(* CODESYS project codesys_webvisu_opcua.project

Project tree, tasks and I/O mapping:
  Device : CODESYS Control for Raspberry Pi SL, CODESYS GmbH, order no. 2302000009, version 4.8.0.0
    application app
      libraries: Standard, 3.5.18.0 (System); Memory, * (3S - Smart Software Solutions GmbH); Util, 3.5.19.0 (System); CmpSysEthernet, 3.4.3.0 (3S - Smart Software Solutions GmbH); VisuDialogs, * (System); CAA Callback Extern, 3.5.17.0 (CAA Technical Workgroup); SysTypes Interfaces, 3.5.2.0 (System); SysMem, 3.5.17.0 (System); CmpErrors Interfaces, * (System); CAA SerialCom, 3.5.17.0 (CAA Technical Workgroup); SysSocket, 3.5.19.0 (System)
      task MainTask (cyclic, interval 4 ms, priority 0) calls MAIN
      task VISU_TASK (cyclic, interval 100 ms, priority 31) calls VisuElems.Visu_Prg
      program MAIN [ST]
      Symbols
      visualisation VISU
      Kommunikationsverwalter
        OPC_UA_Symbols
          Informationsmodell
      function block FB_DEMO [ST]: add2
    SoftMotion General Axis Pool
      x_axis : SM_Drive_Virtual, 3S - Smart Software Solutions GmbH, order no. 1805, version 4.0.0.0
          settings: wDriveID = 0; fSWMaxVelocity = 100000; fSWMaxAcceleration = 100000; fSWMaxDeceleration = 100000; fRampJerk = 1e7; fSWLimitPositive = 3000; fSWLimitNegative = -500; fSWLimitDeceleration = 0.0; fSWErrorMaxDistance = 0.0
      y_axis : SM_Drive_Virtual, 3S - Smart Software Solutions GmbH, order no. 1805, version 4.0.0.0
          settings: fSWMaxVelocity = 100000; fSWMaxAcceleration = 100000; fSWMaxDeceleration = 100000; fRampJerk = 1e7; fSWLimitPositive = 3000; fSWLimitNegative = -3000; fSWLimitDeceleration = 0.0; fSWErrorMaxDistance = 0.0
      z_axis : SM_Drive_Virtual, 3S - Smart Software Solutions GmbH, order no. 1805, version 4.0.0.0
          settings: wDriveID = 2; fSWMaxVelocity = 100000; fSWMaxAcceleration = 100000; fSWMaxDeceleration = 100000; fRampJerk = 1e7; fSWLimitPositive = 100; fSWLimitNegative = -1000; fSWLimitDeceleration = 0.0; fSWErrorMaxDistance = 0.0
      a_axis : SM_Drive_Virtual, 3S - Smart Software Solutions GmbH, order no. 1805, version 4.0.0.0
          settings: wDriveID = 3; fSWMaxVelocity = 100000; fSWMaxAcceleration = 100000; fSWMaxDeceleration = 100000; fRampJerk = 1e7; fSWLimitPositive = 360; fSWLimitNegative = -360; fSWLimitDeceleration = 0.0; fSWErrorMaxDistance = 0.0
      r_axis : SM_Drive_Virtual, 3S - Smart Software Solutions GmbH, order no. 1805, version 4.0.0.0
          settings: wDriveID = 4; fSWMaxVelocity = 100000; fSWMaxAcceleration = 100000; fSWMaxDeceleration = 100000; fRampJerk = 1e7; fSWLimitPositive = 360; fSWLimitNegative = -360; fSWLimitDeceleration = 0.0; fSWErrorMaxDistance = 0.0
    GPIOs_A_B : GPIOs B+/Pi2, 3S - Smart Software Solutions GmbH, version 4.5.0.0
        unmapped channels: digital inputs (GPIO0..GPIO31), digital outputs (GPIO0..GPIO31)
    I²C
    SPI
      SPI_master_CS1 : SPI master, 3S - Smart Software Solutions GmbH, version 1.0.0.0
          settings: SPI port = '/dev/spidev0.1'; _diBitsPerWord = 8; _diMaxSpeed = 2000000
        blp : ABBTS_BLP_V2, ABB Technikerschule, version 1.0
    Onewire
    Camera device
      <Leer>
    Ethernet : Ethernet, 3S - Smart Software Solutions GmbH, version 4.1.0.0
        settings: IPAddress = [127,0,0,1]; SubnetMask = [255,0,0,0]; GatewayAddress = [0,0,0,0]; NetworkInterfaceName = 'lo'; NetworkInterfaceName = "lo"; SaveCommunicationSettings = FALSE
      ModbusTCP_Slave_OLED_Port_503 : ModbusTCP Slave Device, 3S - Smart Software Solutions GmbH, version 4.3.0.0
          settings: Port = 503
          output app.blp.oled.awToOled : ARRAY[0..32] OF WORD  // Ausgänge
          unmapped channels: Eingänge
  libraries: Util, 3.5.19.0 (System)
  text list GlobalTextList
  00000000-0000-0000-0000-000000000000|D:\Dropbox\ABBTS_LABOR_DOZ\LERNPLATTFORM\V2\PCB\_BOM\ADAPTER_RPI_REV3.pdf
  00000000-0000-0000-0000-000000000000|D:\Dropbox\Lernplattformen\01_Basis\SCHEMA_FOTOS\V2\ADAPTER_RPI_REV3.jpg
  00000000-0000-0000-0000-000000000000|D:\Dropbox\ABBTS_LABOR_DOZ\LERNPLATTFORM\V2\PCB\_BOM\DIT_16IN_16_OUT_REV0.pdf
  00000000-0000-0000-0000-000000000000|D:\Dropbox\Lernplattformen\01_Basis\SCHEMA_FOTOS\V2\DIT_16IN_16_OUT_REV0_1.jpg
  00000000-0000-0000-0000-000000000000|D:\Dropbox\ABBTS_LABOR_DOZ\LERNPLATTFORM\V2\PCB\_BOM\IO_LCD_REV2.pdf
  00000000-0000-0000-0000-000000000000|D:\Dropbox\Lernplattformen\01_Basis\SCHEMA_FOTOS\V2\IO_LCD_REV2.jpg
  00000000-0000-0000-0000-000000000000|D:\Dropbox\ABBTS_LABOR_DOZ\LERNPLATTFORM\V2\PCB\_BOM\TRANSFER_TRESOR_REV2.pdf
  00000000-0000-0000-0000-000000000000|D:\Dropbox\Lernplattformen\01_Basis\SCHEMA_FOTOS\V2\TRANSFER_TRESOR_REV2.jpg
*)

// Device/app/MAIN
PROGRAM MAIN
VAR
	rBogenmass: REAL;
	rPi: REAL := 3.14159;
	rMoveX: REAL;
	rRadius: REAL := 50.0;
	rMoveY: REAL;
	rPunktWinkel: REAL;
	arDatenfeld: ARRAY[0..9] OF REAL;
	
	fbDemo: FB_DEMO;
END_VAR

// Rotation eines roten Punktes auf eienm Kreis
rBogenmass := rBogenmass + 0.005;
IF (rBogenmass > (2*rPi)) THEN
	rBogenmass := 0.0;
END_IF
rMoveX := rRadius * COS(rBogenmass);
rMoveY := rRadius * SIN(rBogenmass);
rPunktWinkel := rBogenmass*180.0/rPi;

fbDemo();

(*
https://github.com/FreeOpcUa/opcua-modeler
https://opcua.rocks/custom-information-models/
https://pypi.org/project/opcua-modeler/




*)

END_PROGRAM

// Device/app/FB_DEMO
FUNCTION_BLOCK PUBLIC FB_DEMO
VAR_INPUT
END_VAR
VAR_OUTPUT
END_VAR
VAR
END_VAR

METHOD PUBLIC add2 : REAL
VAR_INPUT
	in1: REAL;
	in2: REAL;
END_VAR
add2 := in1 + in2;
END_METHOD

END_FUNCTION_BLOCK

// Device/app/VISU
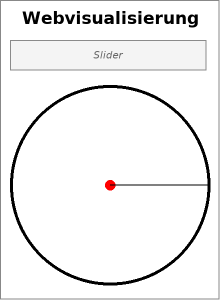
VISUALIZATION VISU  // 220x300
    Ellipse (109,180 2x10)
        p3560616238: MAIN.rMoveX
        p2738717112: MAIN.rMoveY
    Ellipse (10,85 200x200)
    Ellipse (105,180 10x10)
        p3560616238: MAIN.rMoveX
        p2738717112: MAIN.rMoveY
    Line (210,185) (110,185)
        p2858320360: MAIN.rPunktWinkel
    Rectangle (0,0 221x36), "Webvisualisierung"
    Slider (10,40 196x30), variable: MAIN.rRadius, scale 0..100
END_VISUALIZATION
